(* Logix 5000 project; controller PLC_MCC1201_220AP1 vendor 1 type 14 code 164 rev 35.11; software revision 35.00; part 25 of 25 *)
(* tags used below, declared in another part *)
   LEHR_dLehrPositionAdvancement : DINT;
   SnaprollHMW_dOffset_cmm : DINT;
   SnaprollUPS_DistanceFromSnaproll_cmm : DINT;
   TMP_dSnaprollCut_cmm : DINT;
   TMP_xCutOnSnaproll_cmm : BOOL;
   AUX_xInitialize : BOOL;
   GP_NetDiag : GP_NetworkDiag;
   GP_OB_InitializeDiag : GP_OB_Initialize;
   GP_OB_InitializeDiag_STC : GP_OB_Initialize_STC;
   M225 : MAC_EMERGENCYXCUT;
   MCC1201_rgtDiagModule_HMI : GP_NetworkDiag_v1[50];
   N54 : DINT[501];
   TMP_dIndex : DINT;
   Z200 : MAC_Zone_ML;
   Z200_UPS : ZONE_UPS;
   Z200_UPS_HMR : ZONE_UPS_HMR;
(* MainProgram, continued *)

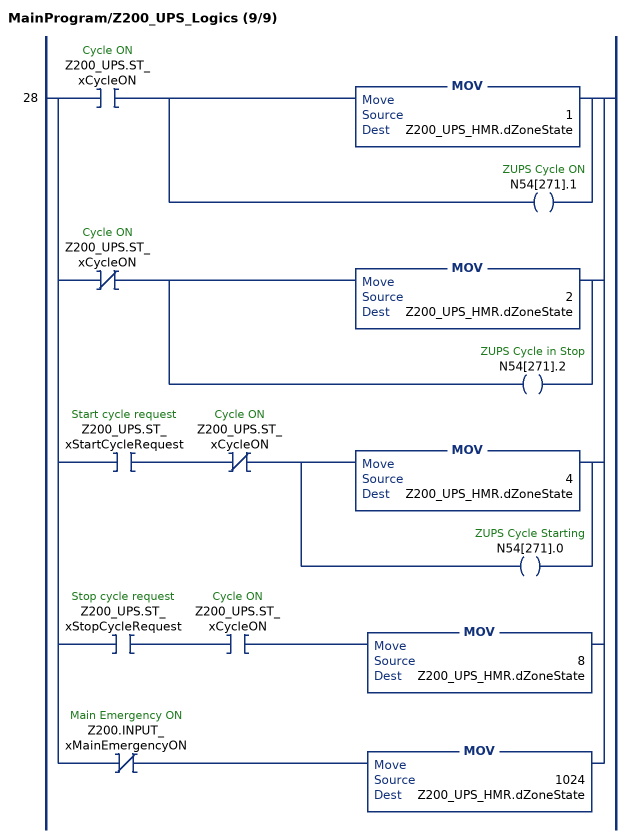
   [picture p437: MainProgram/Z200_UPS_Logics rungs 28-28]
   28: [XIC(Z200_UPS.ST_xCycleON) [MOV(1,Z200_UPS_HMR.dZoneState) ,OTE(N54[271].1) ] ,XIO(Z200_UPS.ST_xCycleON) [MOV(2,Z200_UPS_HMR.dZoneState) ,OTE(N54[271].2) ] ,XIC(Z200_UPS.ST_xStartCycleRequest) XIO(Z200_UPS.ST_xCycleON) [MOV(4,Z200_UPS_HMR.dZoneState) ,OTE(N54[271].0) ] ,XIC(Z200_UPS.ST_xStopCycleRequest) XIC(Z200_UPS.ST_xCycleON) MOV(8,Z200_UPS_HMR.dZoneState) ,XIO(Z200.INPUT_xMainEmergencyON) MOV(1024,Z200_UPS_HMR.dZoneState) ];
END_ROUTINE

ROUTINE ZUPS_Snaproll_SearchCut   (* structured text *)
   TMP_xCutOnSnaproll_cmm := 0;
   FOR TMP_dIndex:=0 to M225.AUX_dTankElementCounter do
   	TMP_dSnaprollCut_cmm := LEHR_dLehrPositionAdvancement + SnaprollUPS_DistanceFromSnaproll_cmm - M225.AUX_rgdCutTank[TMP_dIndex] - SnaprollHMW_dOffset_cmm;
   	IF TMP_dSnaprollCut_cmm > 0 AND TMP_dSnaprollCut_cmm < 30000 then
   		TMP_xCutOnSnaproll_cmm:=1;
   	END_IF;
   END_FOR;
END_ROUTINE
END_PROGRAM

PROGRAM Modules   (* main routine Main *)

ROUTINE Main   (* ladder *)
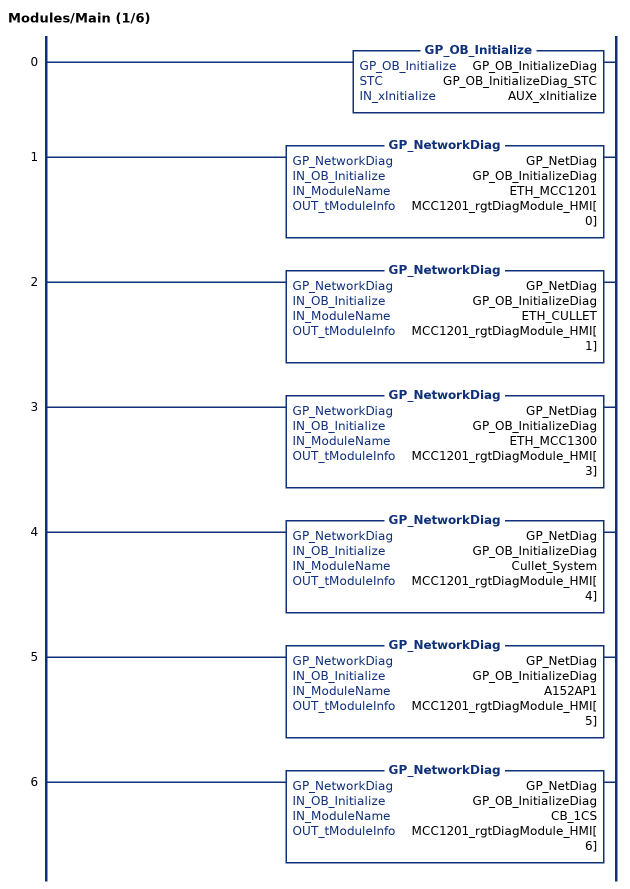
   0: GP_OB_Initialize(GP_OB_InitializeDiag,GP_OB_InitializeDiag_STC,AUX_xInitialize);
   1: GP_NetworkDiag(GP_NetDiag,GP_OB_InitializeDiag,ETH_MCC1201,MCC1201_rgtDiagModule_HMI[0]);
   2: GP_NetworkDiag(GP_NetDiag,GP_OB_InitializeDiag,ETH_CULLET,MCC1201_rgtDiagModule_HMI[1]);
   3: GP_NetworkDiag(GP_NetDiag,GP_OB_InitializeDiag,ETH_MCC1300,MCC1201_rgtDiagModule_HMI[3]);
   4: GP_NetworkDiag(GP_NetDiag,GP_OB_InitializeDiag,Cullet_System,MCC1201_rgtDiagModule_HMI[4]);
   5: GP_NetworkDiag(GP_NetDiag,GP_OB_InitializeDiag,A152AP1,MCC1201_rgtDiagModule_HMI[5]);
   6: GP_NetworkDiag(GP_NetDiag,GP_OB_InitializeDiag,CB_1CS,MCC1201_rgtDiagModule_HMI[6]);
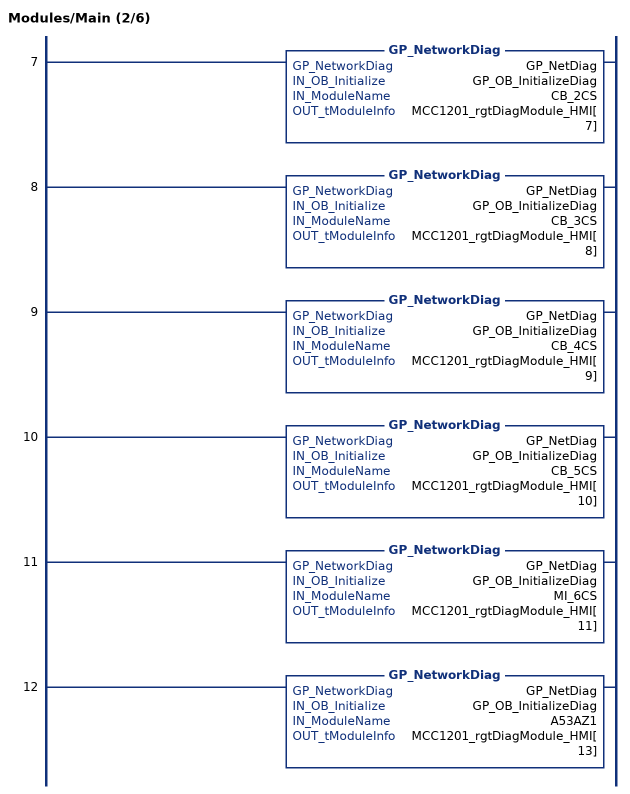
   7: GP_NetworkDiag(GP_NetDiag,GP_OB_InitializeDiag,CB_2CS,MCC1201_rgtDiagModule_HMI[7]);
   8: GP_NetworkDiag(GP_NetDiag,GP_OB_InitializeDiag,CB_3CS,MCC1201_rgtDiagModule_HMI[8]);
   9: GP_NetworkDiag(GP_NetDiag,GP_OB_InitializeDiag,CB_4CS,MCC1201_rgtDiagModule_HMI[9]);
   10: GP_NetworkDiag(GP_NetDiag,GP_OB_InitializeDiag,CB_5CS,MCC1201_rgtDiagModule_HMI[10]);
   11: GP_NetworkDiag(GP_NetDiag,GP_OB_InitializeDiag,MI_6CS,MCC1201_rgtDiagModule_HMI[11]);
   12: GP_NetworkDiag(GP_NetDiag,GP_OB_InitializeDiag,A53AZ1,MCC1201_rgtDiagModule_HMI[13]);
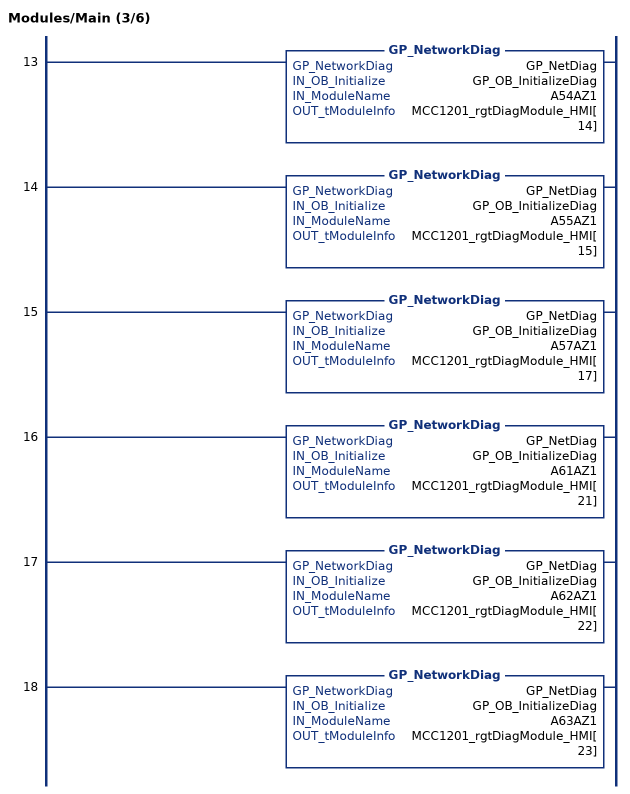
   13: GP_NetworkDiag(GP_NetDiag,GP_OB_InitializeDiag,A54AZ1,MCC1201_rgtDiagModule_HMI[14]);
   14: GP_NetworkDiag(GP_NetDiag,GP_OB_InitializeDiag,A55AZ1,MCC1201_rgtDiagModule_HMI[15]);
   15: GP_NetworkDiag(GP_NetDiag,GP_OB_InitializeDiag,A57AZ1,MCC1201_rgtDiagModule_HMI[17]);
   16: GP_NetworkDiag(GP_NetDiag,GP_OB_InitializeDiag,A61AZ1,MCC1201_rgtDiagModule_HMI[21]);
   17: GP_NetworkDiag(GP_NetDiag,GP_OB_InitializeDiag,A62AZ1,MCC1201_rgtDiagModule_HMI[22]);
   18: GP_NetworkDiag(GP_NetDiag,GP_OB_InitializeDiag,A63AZ1,MCC1201_rgtDiagModule_HMI[23]);
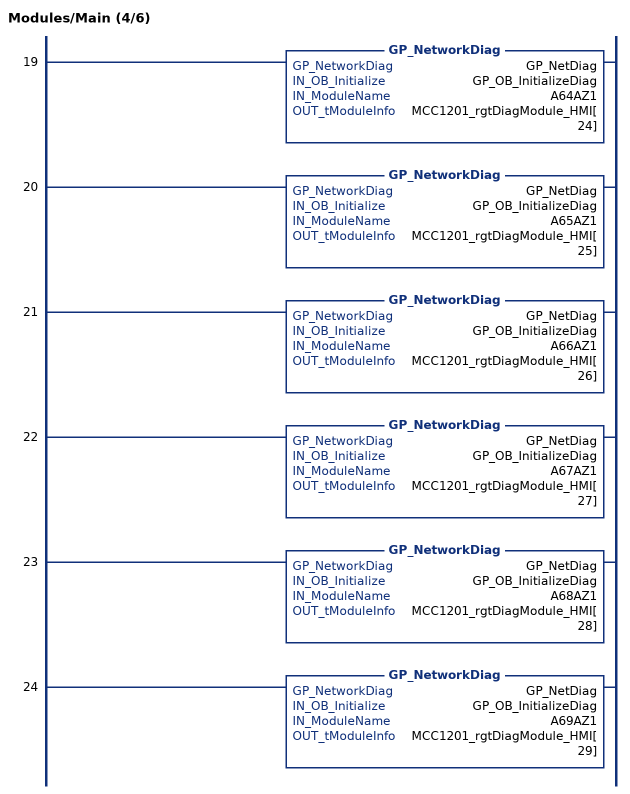
   19: GP_NetworkDiag(GP_NetDiag,GP_OB_InitializeDiag,A64AZ1,MCC1201_rgtDiagModule_HMI[24]);
   20: GP_NetworkDiag(GP_NetDiag,GP_OB_InitializeDiag,A65AZ1,MCC1201_rgtDiagModule_HMI[25]);
   21: GP_NetworkDiag(GP_NetDiag,GP_OB_InitializeDiag,A66AZ1,MCC1201_rgtDiagModule_HMI[26]);
   22: GP_NetworkDiag(GP_NetDiag,GP_OB_InitializeDiag,A67AZ1,MCC1201_rgtDiagModule_HMI[27]);
   23: GP_NetworkDiag(GP_NetDiag,GP_OB_InitializeDiag,A68AZ1,MCC1201_rgtDiagModule_HMI[28]);
   24: GP_NetworkDiag(GP_NetDiag,GP_OB_InitializeDiag,A69AZ1,MCC1201_rgtDiagModule_HMI[29]);
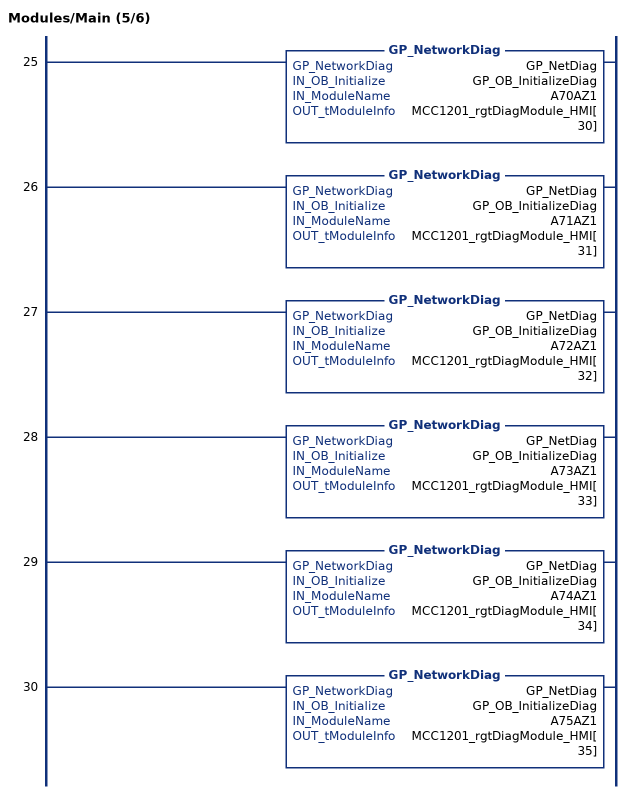
   25: GP_NetworkDiag(GP_NetDiag,GP_OB_InitializeDiag,A70AZ1,MCC1201_rgtDiagModule_HMI[30]);
   26: GP_NetworkDiag(GP_NetDiag,GP_OB_InitializeDiag,A71AZ1,MCC1201_rgtDiagModule_HMI[31]);
   27: GP_NetworkDiag(GP_NetDiag,GP_OB_InitializeDiag,A72AZ1,MCC1201_rgtDiagModule_HMI[32]);
   28: GP_NetworkDiag(GP_NetDiag,GP_OB_InitializeDiag,A73AZ1,MCC1201_rgtDiagModule_HMI[33]);
   29: GP_NetworkDiag(GP_NetDiag,GP_OB_InitializeDiag,A74AZ1,MCC1201_rgtDiagModule_HMI[34]);
   30: GP_NetworkDiag(GP_NetDiag,GP_OB_InitializeDiag,A75AZ1,MCC1201_rgtDiagModule_HMI[35]);
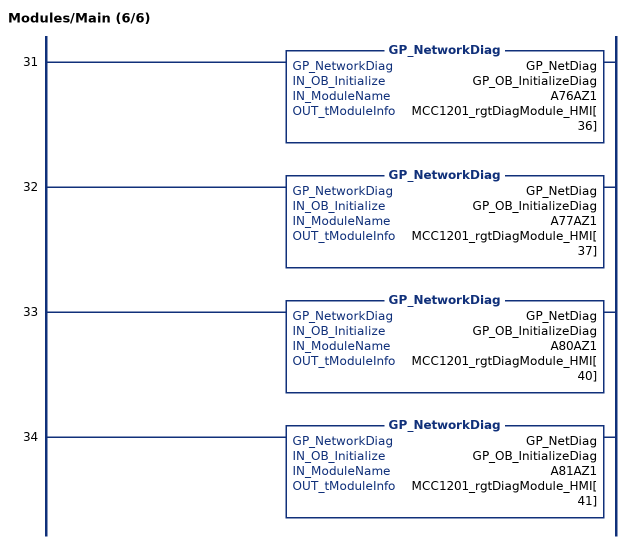
   31: GP_NetworkDiag(GP_NetDiag,GP_OB_InitializeDiag,A76AZ1,MCC1201_rgtDiagModule_HMI[36]);
   32: GP_NetworkDiag(GP_NetDiag,GP_OB_InitializeDiag,A77AZ1,MCC1201_rgtDiagModule_HMI[37]);
   33: GP_NetworkDiag(GP_NetDiag,GP_OB_InitializeDiag,A80AZ1,MCC1201_rgtDiagModule_HMI[40]);
   34: GP_NetworkDiag(GP_NetDiag,GP_OB_InitializeDiag,A81AZ1,MCC1201_rgtDiagModule_HMI[41]);
END_ROUTINE
END_PROGRAM
